screen "tryb_manualny" 800x480
   on GenerateScreen: SetTag("Tag_ScreenNumber", 2)
   TextField "Text field_1" at 282,4 size 223x34; Text 'TRYB MANUALNY'
   TextField "Text field_4" at 512,155 size 171x61; Text 'STOPIEŃ OTWARCIA OKIEN OTWIERANIE OKIEN'
   Button "Button_4" at 518,261 size 80x70; TextOff 'PODLEWANIE'
      on Click: InvertBit("Przycisk_podlewania_manual")
   Button "Button_5" at 611,261 size 80x70; TextOff 'GRZANIE'
      on Click: InvertBit("Przycisk_grzanie_manual")
   Button "Button_6" at 701,261 size 80x70; TextOff 'WENTYLACJA'
      on Click: InvertBit("Przycisk_wentylacja_manual")
   GraphicView "Graphic view_1" at 710,356 size 60x60; Picture "fan_4829316"
      Visibility <- "Wentylator"
   GraphicView "Graphic view_6" at 622,356 size 60x60; Picture "heater_4463010"
      Visibility <- "Grzałka"
   GraphicView "Graphic view_7" at 527,356 size 64x60; Picture "irrigation_18631825"
      Visibility <- "Pompa_podlewanie"
   GraphicView "Graphic view_9" at 710,356 size 60x60; Picture "fan_off"
      Visibility <- "Wentylator"
   GraphicView "Graphic view_10" at 622,356 size 60x60; Picture "heater_off"
      Visibility <- "Grzałka"
   GraphicView "Graphic view_11" at 527,356 size 64x60; Picture "irrigation_off"
      Visibility <- "Pompa_podlewanie"
   Button "Button_14" at 3,1 size 43x43; TextOff 'DOM'; PictureOff "home_1"
      on Click: ActivateScreen("Root screen", 0)
   Button "Button_1" at 750,0 size 50x50; TextOff 'Text'; PictureOff "Back_arrow"
      on Click: function_efd93a16()
   Circle "Circle_1" at 541,428 size 42x42
      Visibility <- "Pompa_podlewanie"
   Circle "Circle_4" at 541,428 size 42x42
      Visibility <- "Pompa_podlewanie"
   Circle "Circle_2" at 631,428 size 42x42
      Visibility <- "Grzałka"
   Circle "Circle_5" at 631,428 size 42x42
      Visibility <- "Grzałka"
   Circle "Circle_3" at 720,428 size 41x41
      Visibility <- "Wentylator"
   Circle "Circle_6" at 720,428 size 41x41
      Visibility <- "Wentylator"
   TextField "Text field_8" at 405,71 size 117x61; Text 'STOPIEŃ OTWARCIA OKIEN STOPIEŃ ZASŁONIECIA ROLET'
   Bar "Bar_6" at 625,71 size 165x66; MinimumValue 0; MaximumValue 100
      ProcessValue <- "Stopien_zasloniecia_rolet_manual"
   Button "Button_3" at 532,109 size 80x50; TextOff '+ / ODSŁOŃ'
      on Click: function_b9b71300("Stopien_zasloniecia_rolet_manual", 5)
   Button "Button_7" at 530,49 size 80x50; TextOff '- / ZASŁOŃ'
      on Press: function_dd21b452("Stopien_zasloniecia_rolet_manual", 5)
   Button "Button_2" at 425,261 size 80x70; TextOff 'PODLEWANIE / MIKROZRASZANIE'
      on Click: InvertBit("Przycisk_zraszania_manual")
   GraphicView "Graphic view_2" at 434,356 size 60x60; Picture "sprinkler_4552152"
      Visibility <- "Pompa_zraszacze"
   GraphicView "Graphic view_3" at 434,356 size 60x60; Picture "sprinkler"
      Visibility <- "Pompa_zraszacze"
   Circle "Circle_7" at 443,428 size 42x42
      Visibility <- "Pompa_zraszacze"
   Circle "Circle_8" at 443,428 size 42x42
      Visibility <- "Pompa_zraszacze"
   Switch "Switch_1" at 499,199 size 209x37; CaptionText 'Switch'; TextOff 'ZAMKNIĘTE'; TextOn 'OTWARTE'
      ProcessValue <- "Otwarcie_okien_man"
   TextField "Text field_3" at 10,365 size 166x23; Text 'SZYBKOŚĆ WIATRU'
   IOField "I/O field_3" at 61,397 size 70x65; FormatPattern 999
      ProcessValue <- "Czujnik_wiatru"
   IOField "I/O field_1" at 47,179 size 101x32; FormatPattern 99999
      ProcessValue <- "Czujnik_natezenia_światła"
   TextField "Text field_15" at 128,398 size 52x72; Text 'Km h'
   IOField "I/O field_2" at 43,282 size 83x65; FormatPattern 9999
      ProcessValue <- "Wewnetrzny_czujnik_CO2"
   TextField "Text field_11" at 117,291 size 69x39; Text 'ppm'
   TextField "Text field_5" at 13,138 size 204x23; Text 'INSOLATION / NASŁONECZNIENIE / SONNENEINSTRAHLUNG'
   IOField "I/O field_8" at 57,85 size 93x40; FormatPattern 99.99
      ProcessValue <- "Temperatura_wewnetrzna"
   TextField "Text field_20" at 26,42 size 137x42; Text 'TEMPERATURA TEMPERATURA WEWNTĘTRZNA'
   TextField "Text field_7" at 199,365 size 175x23; Text 'WILGOTNOŚĆ GLEBY'
   IOField "I/O field_5" at 247,283 size 83x65; FormatPattern 9999
      ProcessValue <- "Zewnetrzny_czujnik_CO2"
   IOField "I/O field_4" at 265,164 size 69x65; FormatPattern 999
      ProcessValue <- "Czujnik_wilgotności_powietrza"
   IOField "I/O field_6" at 260,395 size 68x65; FormatPattern 999
      ProcessValue <- "Czujnik_wilgotności_gleby"
   TextField "Text field_12" at 323,172 size 47x46; Text '%'
   TextField "Text field_13" at 320,406 size 47x46; Text '%'
   TextField "Text field_16" at 326,292 size 69x39; Text 'ppm'
   IOField "I/O field_9" at 247,75 size 97x65; FormatPattern 99.99
      ProcessValue <- "Temperatura_zewnetrzna"
   TextField "Text field_23" at 332,80 size 46x46; Text '°C'
   TextField "Text field_22" at 227,43 size 132x42; Text 'TEMPERATURA TEMPERATURA ZEWNĘTRZNA'
   TextField "Text field_9" at 228,246 size 123x42; Text 'STĘŻENIE CO2 ZEWNĘTRZNE STĘŻENIE CO2'
   TextField "Text field_6" at 180,137 size 223x42; Text 'WILGOTNOŚĆ POWIETRZA WILGOTNOŚĆ POWIETRZA'
   TextField "Text field_14" at 139,160 size 47x72; Text 'W m²'
   TextField "Text field_21" at 140,80 size 46x46; Text '°C'
   GraphicView "Graphic view_4" at 419,176 size 60x60; Picture "window_11250237"
   GraphicView "Graphic view_5" at 196,172 size 50x50; Picture "sensor_4212519"
   GraphicView "Graphic view_8" at 3,172 size 50x50; Picture "sensor_4212513"
   GraphicView "Graphic view_12" at 2,77 size 50x50; Picture "Thermometer_icon"
   GraphicView "Graphic view_13" at 198,77 size 50x50; Picture "Thermometer_icon"
   GraphicView "Graphic view_14" at 2,292 size 40x40; Picture "sensor_2828470"
   GraphicView "Graphic view_15" at 196,290 size 40x40; Picture "sensor_2828470"
   GraphicView "Graphic view_16" at 197,402 size 50x50; Picture "soil-sensor_11298794"
   GraphicView "Graphic view_17" at 2,406 size 50x50; Picture "anemometer_1113716"
   TextField "Text field_2" at 26,246 size 124x42; Text 'STĘŻENIE CO2 WEWNĘTRZNE STĘŻENIE CO2'

screen "praca" 800x480
   on GenerateScreen: SetTag("Tag_ScreenNumber", 5)
   GraphicView "Graphic view_4" at 274,396 size 70x70; Picture "soil-sensor_11298794"
   GraphicView "Graphic view_3" at 3,175 size 70x70; Picture "sensor_4212513"
   GraphicView "Graphic view_5" at 267,175 size 70x70; Picture "sensor_4212519"
   GraphicView "Graphic view_1" at 559,396 size 70x70; Picture "fan_4829316"
      Visibility <- "Wentylator"
   GraphicView "Graphic view_6" at 560,270 size 70x70; Picture "heater_4463010"
      Visibility <- "Grzałka"
   GraphicView "Graphic view_7" at 559,164 size 70x70; Picture "irrigation_18631825"
      Visibility <- "Pompa_podlewanie"
   GraphicView "Graphic view_8" at 11,397 size 70x70; Picture "anemometer_1113716"
   GraphicView "Graphic view_9" at 559,396 size 70x70; Picture "fan_off"
      Visibility <- "Wentylator"
   GraphicView "Graphic view_10" at 560,270 size 70x70; Picture "heater_off"
      Visibility <- "Grzałka"
   GraphicView "Graphic view_11" at 559,164 size 70x70; Picture "irrigation_off"
      Visibility <- "Pompa_podlewanie"
   GraphicView "Graphic view_12" at 278,267 size 70x70; Picture "sensor_2828470"
   TextField "Text field_1" at 52,152 size 204x23; Text 'INSOLATION / NASŁONECZNIENIE / SONNENEINSTRAHLUNG'
   TextField "Text field_3" at 44,373 size 166x23; Text 'SZYBKOŚĆ WIATRU'
   TextField "Text field_5" at 289,152 size 223x23; Text 'WILGOTNOŚĆ POWIETRZA'
   TextField "Text field_6" at 318,373 size 175x23; Text 'WILGOTNOŚĆ GLEBY'
   TextField "Text field_7" at 628,148 size 116x23; Text 'PODLEWANIE'
   TextField "Text field_8" at 638,252 size 80x23; Text 'GRZANIE'
   TextField "Text field_9" at 627,373 size 117x23; Text 'WENTYLACJA'
   TextField "Text field_10" at 81,3 size 256x34; Text 'PODGLĄD NA ŻYWO'
   Button "Button_1" at 750,0 size 50x50; TextOff 'WRÓĆ'; PictureOff "Back_arrow"
      on Click: function_efd93a16(); SetBit("HMI_Reset_Trybow")
   Button "Button_2" at 3,1 size 43x43; TextOff 'DOM'; PictureOff "home_1"
      on Click: ActivateScreen("Root screen", 0); SetBit("HMI_Reset_Trybow")
   IOField "I/O field_3" at 94,402 size 70x65; FormatPattern 999
      ProcessValue <- "Czujnik_wiatru"
   IOField "I/O field_5" at 348,277 size 83x65; FormatPattern 9999
      ProcessValue <- "Zewnetrzny_czujnik_CO2"
   IOField "I/O field_4" at 377,172 size 69x65; FormatPattern 999
      ProcessValue <- "Czujnik_wilgotności_powietrza"
   IOField "I/O field_6" at 381,397 size 68x65; FormatPattern 999
      ProcessValue <- "Czujnik_wilgotności_gleby"
   TextField "Text field_12" at 446,190 size 47x46; Text '%'
   TextField "Text field_13" at 466,405 size 47x46; Text '%'
   TextField "Text field_14" at 192,164 size 47x72; Text 'W m²'
   IOField "I/O field_1" at 83,190 size 101x32; FormatPattern 99999
      ProcessValue <- "Czujnik_natezenia_światła"
   TextField "Text field_15" at 173,402 size 52x72; Text 'Km h'
   Circle "Circle_1" at 703,188 size 48x48
      Visibility <- "Pompa_podlewanie"
   Circle "Circle_2" at 702,283 size 48x48
      Visibility <- "Grzałka"
   TextField "Text field_16" at 447,283 size 69x39; Text 'ppm'
   Circle "Circle_4" at 703,188 size 48x48
      Visibility <- "Pompa_podlewanie"
   Circle "Circle_5" at 702,283 size 48x48
      Visibility <- "Grzałka"
   Circle "Circle_3" at 703,415 size 48x48
      Visibility <- "Wentylator"
   Circle "Circle_6" at 703,415 size 48x48
      Visibility <- "Wentylator"
   TextField "Text field_17" at 381,3 size 288x34; Text 'PODGLĄD NA ŻYWO / TRYB AUTOMATYCZNY'
      Visibility <- "HMI_Aktywacja_trybu_automatycznego"
   GraphicView "Graphic view_13" at 560,63 size 70x70; Picture "sprinkler_4552152"
      Visibility <- "Pompa_zraszacze"
   GraphicView "Graphic view_14" at 560,63 size 70x70; Picture "sprinkler"
      Visibility <- "Pompa_zraszacze"
   Circle "Circle_7" at 703,83 size 48x48
      Visibility <- "Pompa_zraszacze"
   Circle "Circle_8" at 703,83 size 48x48
      Visibility <- "Pompa_zraszacze"
   TextField "Text field_19" at 609,44 size 156x23; Text 'PODLEWANIE / MIKROZRASZANIE'
   GraphicView "Graphic view_15" at 0,66 size 70x70; Picture "Thermometer_icon"
   IOField "I/O field_8" at 73,73 size 97x65; FormatPattern 99.99
      ProcessValue <- "Temperatura_wewnetrzna"
   TextField "Text field_21" at 171,85 size 46x46; Text '°C'
   GraphicView "Graphic view_16" at 275,66 size 70x70; Picture "Thermometer_icon"
   IOField "I/O field_9" at 348,73 size 97x65; FormatPattern 99.99
      ProcessValue <- "Temperatura_zewnetrzna"
   TextField "Text field_23" at 447,82 size 46x46; Text '°C'
   TextField "Text field_20" at 57,44 size 137x42; Text 'TEMPERATURA TEMPERATURA WEWNTĘTRZNA'
   TextField "Text field_22" at 334,44 size 132x42; Text 'TEMPERATURA TEMPERATURA ZEWNĘTRZNA'
   GraphicView "Graphic view_2" at 11,273 size 70x70; Picture "sensor_2828470"
   IOField "I/O field_2" at 81,283 size 83x65; FormatPattern 9999
      ProcessValue <- "Wewnetrzny_czujnik_CO2"
   TextField "Text field_11" at 180,289 size 69x39; Text 'ppm'
   TextField "Text field_2" at 83,252 size 124x42; Text 'STĘŻENIE CO2 WEWNĘTRZNE STĘŻENIE CO2'
   TextField "Text field_4" at 352,256 size 123x42; Text 'STĘŻENIE CO2 ZEWNĘTRZNE STĘŻENIE CO2'
   TextField "Text field_18" at 381,3 size 211x34; Text 'TRYB RECEPTUR'
      Visibility <- "HMI_Aktywacja_trybu_Receptur"

Template "Template_1" 800x480
   Button "Exit" at 671,429 size 71x50; TextOn 'Exit'; TextOff 'Exit'; PictureOn "ExitRuntime_KTP700_Basic_PN_TR"; PictureOff "ExitRuntime_KTP700_Basic_PN_TR"
      on Release: StopRuntime(0)
   Button "Alarms" at 524,429 size 71x50; TextOn 'Alarms'; TextOff 'Alarms'; PictureOn "AlarmDisplay_KTP700_Basic_PN_TR"; PictureOff "AlarmDisplay_KTP700_Basic_PN_TR"
      on Release: function_ef3f5d25("Alarm window_Unacknowledged", -1)
   Button "Start screen" at 169,429 size 71x50; TextOn 'Start screen'; TextOff 'Start screen'; PictureOn "NavigateHome_KTP700_Basic_PN_TR"; PictureOff "NavigateHome_KTP700_Basic_PN_TR"
      on Release: ActivateScreen("Root screen", 0)
      Visibility <- "AlwaysTRUE"
   Button "Language" at 377,429 size 71x50; TextOn 'Language'; TextOff 'Language'; PictureOn "ToggleLanguage_KTP700_Basic_PN_TR"; PictureOff "ToggleLanguage_KTP700_Basic_PN_TR"
      on Release: function_fb9197e8(-1)

screen "Receptury" 800x480
   RecipeView "Recipe view_1" at 0,38 size 799x413; Recipe "Receptura_nr1"; RecipeNameCaption 'Recipe Name: / Wybierz Recepturę / Rezepturname:'; EntryNameCaption 'Entry Name / Zapisane Parametry / Eintragsname'; DataRecordNameCaption 'Data Record Name: / Wybierz Recepturę / Datensatzname:'
   GraphicView "Graphic view_1" at 529,152 size 35x35; Picture "Thermometer_icon"
   GraphicView "Graphic view_2" at 529,190 size 35x35; Picture "sensor_4212519"
   GraphicView "Graphic view_3" at 529,230 size 35x35; Picture "soil-sensor_11298794"
   GraphicView "Graphic view_4" at 529,269 size 35x35; Picture "window_11250237"
   GraphicView "Graphic view_5" at 529,308 size 35x35; Picture "sensor_2828470"
   GraphicView "Graphic view_6" at 529,348 size 35x35; Picture "sensor_4212513"
   TextField "Text field_11" at 569,150 size 39x38; Text '°C'
   TextField "Text field_18" at 569,190 size 39x38; Text '%'
   TextField "Text field_1" at 569,230 size 39x38; Text '%'
   TextField "Text field_2" at 564,269 size 57x32; Text '1/0'
   TextField "Text field_16" at 563,308 size 55x32; Text 'ppm'
   TextField "Text field_6" at 576,339 size 28x50; Text '°C W m'
   TextField "Text field_3" at 593,362 size 31x17; Text '2'
   Button "Button_1" at 750,0 size 50x50; TextOff 'WRÓĆ'; PictureOff "Back_arrow"
      on Click: function_efd93a16()
   Button "Button_14" at 3,1 size 43x43; TextOff 'DOM'; PictureOff "home_1"
      on Click: ActivateScreen("Root screen", 0)
   TextField "Text field_4" at 320,2 size 170x37; Text 'RECEPTURY'
   TextField "Text field_5" at 12,448 size 50x23; Text 'Nowy'
   TextField "Text field_7" at 69,448 size 57x23; Text 'Zapisz'
   TextField "Text field_8" at 137,448 size 45x23; Text 'Usuń'
   TextField "Text field_9" at 190,438 size 60x42; Text 'Zmień Nazwę'
   TextField "Text field_10" at 663,438 size 66x42; Text 'Załaduj z PLC'
   TextField "Text field_12" at 729,438 size 66x42; Text 'Załaduj do PLC'
   Button "Button_2" at 405,402 size 255x40; TextOff 'ZATWIERDŹ'
      on Click: ResetBit("HMI_Reset_Trybow"); ActivateScreen("praca", 0); SetBit("HMI_Aktywacja_trybu_Receptur")
   TextField "Text field_13" at 456,450 size 173x23; Text 'Przejdź w tryb pracy'
   Button "Button_3" at 256,401 size 140x40; TextOff 'Z'
      on Click: function_ea909784(1, U 0, '\USB_X60.1\record.csv', 2, 1, N)
   TextField "Text field_14" at 266,438 size 113x42; Text 'Zapisz Kopię zapasową'

screen "Symulacja_czujnikow" 800x480
   TextField "Text field_1" at 21,47 size 252x23; Text 'Czujnik Wilgotności powietrza'
   TextField "Text field_2" at 308,47 size 214x23; Text 'Czujnik Wilgotności gleby'
   TextField "Text field_3" at 32,202 size 202x23; Text 'Termometr wewnętrzny'
   TextField "Text field_4" at 323,202 size 197x23; Text 'Termometr zewnętrzny'
   TextField "Text field_5" at 569,47 size 216x23; Text 'Czujnik natężenia światła'
   TextField "Text field_6" at 607,202 size 124x23; Text 'Czujnik wiatru'
   TextField "Text field_7" at 27,346 size 208x23; Text 'Wewnętrzny czujnik CO2'
   TextField "Text field_8" at 306,346 size 202x23; Text 'Zewnętrzny czujnik CO2'
   TextField "Text field_9" at 569,346 size 206x23; Text 'Stopień zasłonięcia rolet'
   IOField "I/O field_4" at 599,83 size 150x60; FormatPattern 9999
      ProcessValue <- "Czujnik_natezenia_światła"
   IOField "I/O field_5" at 599,242 size 150x60; FormatPattern 999
      ProcessValue <- "Czujnik_wiatru"
   IOField "I/O field_6" at 69,375 size 150x60; FormatPattern 9999
      ProcessValue <- "Wewnetrzny_czujnik_CO2"
   IOField "I/O field_7" at 346,375 size 150x60; FormatPattern 9999
      ProcessValue <- "Zewnetrzny_czujnik_CO2"
   IOField "I/O field_8" at 599,375 size 150x60; FormatPattern 999
      ProcessValue <- "Stopien_zasloniecia_rolet"
   IOField "I/O field_10" at 69,83 size 150x60; FormatPattern 999
      ProcessValue <- "Czujnik_wilgotności_powietrza"
   IOField "I/O field_11" at 346,83 size 150x60; FormatPattern 999
      ProcessValue <- "Czujnik_wilgotności_gleby"
   IOField "I/O field_12" at 69,242 size 150x60; FormatPattern 99.9
      ProcessValue <- "Temperatura_wewnetrzna"
   IOField "I/O field_13" at 346,242 size 150x60; FormatPattern 99.9
      ProcessValue <- "Temperatura_zewnetrzna"
   TextField "Text field_10" at 248,5 size 321x34; Text 'ZAPISZ RECEPTURE / SYMULACJA CZUJNIKÓW'
   Button "Button_1" at 750,0 size 50x50; TextOff 'WRÓĆ'; PictureOff "Back_arrow"
      on Click: function_efd93a16()
   Button "Button_14" at 3,1 size 43x43; TextOff 'DOM'; PictureOff "home_1"
      on Click: ActivateScreen("Root screen", 0)

screen "tryb_automatyczny" 800x480
   on GenerateScreen: SetTag("Tag_ScreenNumber", 1)
   IOField "I/O field_1" at 67,301 size 57x40; FormatPattern 99.9
      ProcessValue <- "Temperatura_wewnetrzna"
   Button "Button_1" at 750,0 size 50x50; TextOff 'WRÓĆ'; PictureOff "Back_arrow"
      on Click: function_efd93a16()
   Button "Button_2" at 530,382 size 259x89; TextOff 'ZATWIERDŹ'
      on Click: ResetBit("HMI_Reset_Trybow"); SetBit("HMI_Aktywacja_trybu_automatycznego"); ActivateScreen("praca", 0)
   Bar "Bar_1" at 7,89 size 50x250; MinimumValue 0; MaximumValue 45
      ProcessValue <- "Temperatura_auto"
   TextField "Text field_2" at 1,50 size 132x23; Text 'TEMPERATURA'
   Bar "Bar_2" at 170,90 size 50x250; MinimumValue 0; MaximumValue 100
      ProcessValue <- "Wilgotnosc_powietrza_auto"
   TextField "Text field_3" at 165,47 size 122x42; Text 'WOLGOTNOŚĆ POWIETRZA WILGOTNOŚĆ POWIETRZA'
   Button "Button_3" at 71,94 size 75x45; TextOff '+ / +0.5 °C'
      on Press: function_dd21b452("Temperatura_auto", 0.5)
   Button "Button_7" at 71,162 size 75x45; TextOff '- / -0.5 °C'
      on Press: function_b9b71300("Temperatura_auto", 0.5)
   IOField "I/O field_2" at 67,230 size 62x40; FormatPattern 99.9
      ProcessValue <- "Temperatura_auto"
   TextField "Text field_11" at 122,239 size 23x22; Text '°C'
   TextField "Text field_9" at 122,312 size 23x22; Text '°C'
   Bar "Bar_4" at 335,90 size 50x250; MinimumValue 0; MaximumValue 100
      ProcessValue <- "Wilgotnosc_gleby_auto"
   TextField "Text field_10" at 327,46 size 122x42; Text 'WOLGOTNOŚĆ GLEBY WILGOTNOŚĆ GLEBY'
   Button "Button_8" at 398,111 size 65x40; TextOff '+ / +2%'
      on Click: function_dd21b452("Wilgotnosc_gleby_auto", 2)
   Button "Button_9" at 398,160 size 65x40; TextOff '- / -2%'
      on Click: function_b9b71300("Wilgotnosc_gleby_auto", 2)
   IOField "I/O field_5" at 402,234 size 60x40; FormatPattern 999
      ProcessValue <- "Wilgotnosc_gleby_auto"
   IOField "I/O field_6" at 404,304 size 58x40; FormatPattern 999
      ProcessValue <- "Czujnik_wilgotności_gleby"
   TextField "Text field_12" at 385,222 size 101x22; Text 'USTAWIONA'
   TextField "Text field_13" at 389,293 size 86x22; Text 'AKTUALNA'
   TextField "Text field_14" at 439,243 size 23x22; Text '%'
   TextField "Text field_15" at 439,314 size 23x22; Text '%'
   Button "Button_10" at 229,105 size 65x40; TextOff '+ / +5%'
      on Click: function_dd21b452("Wilgotnosc_powietrza_auto", 5)
   Button "Button_11" at 229,165 size 65x40; TextOff '- / -5%'
      on Click: function_b9b71300("Wilgotnosc_powietrza_auto", 5)
   IOField "I/O field_4" at 234,227 size 66x40; FormatPattern 999
      ProcessValue <- "Wilgotnosc_powietrza_auto"
   IOField "I/O field_7" at 236,299 size 62x40; FormatPattern 999
      ProcessValue <- "Czujnik_wilgotności_powietrza"
   TextField "Text field_16" at 223,214 size 101x22; Text 'USTAWIONA'
   TextField "Text field_17" at 223,285 size 86x22; Text 'AKTUALNA'
   TextField "Text field_18" at 275,236 size 23x22; Text '%'
   TextField "Text field_19" at 275,307 size 23x22; Text '%'
   Button "Button_14" at 3,1 size 43x43; TextOff 'DOM'; PictureOff "home_1"
      on Click: ActivateScreen("Root screen", 0)
   TextField "Text field_4" at 124,384 size 128x23; Text 'SYSTEM OKIEN'
   Switch "Switch_1" at 106,410 size 181x46; TextOn 'ON'; CaptionText 'Switch'; TextOff 'OFF'
      ProcessValue <- "System_okien_auto"
   GraphicView "Graphic view_1" at 128,46 size 40x40; Picture "Thermometer_icon"
   GraphicView "Graphic view_2" at 281,47 size 40x40; Picture "sensor_4212519"
   TextField "Text field_5" at 60,288 size 86x22; Text 'AKTUALNA'
   TextField "Text field_6" at 57,216 size 101x22; Text 'USTAWIONA'
   GraphicView "Graphic view_3" at 443,50 size 40x40; Picture "soil-sensor_11298794"
   TextField "Text field_1" at 250,4 size 288x34; Text 'TRYB AUTOMATYCZNY'
   Bar "Bar_3" at 496,90 size 50x250; MinimumValue 0; MaximumValue 1500
      ProcessValue <- "Naslonecznienie_auto"
   TextField "Text field_7" at 487,38 size 154x40; Text 'WOLGOTNOŚĆ GLEBY NASŁONECZNIENIE'
   GraphicView "Graphic view_4" at 585,65 size 40x40; Picture "sensor_4212513"
   Button "Button_4" at 553,110 size 82x43; TextOff '+ +50 W m'
      on Click: function_dd21b452("Naslonecznienie_auto", 50)
   Button "Button_5" at 554,165 size 82x43; TextOff '- -50 W m'
      on Click: function_b9b71300("Naslonecznienie_auto", 50)
   IOField "I/O field_3" at 561,233 size 61x40; FormatPattern 9999
      ProcessValue <- "Naslonecznienie_auto"
   TextField "Text field_8" at 545,221 size 101x22; Text 'USTAWIONA / USTAWIONE'
   IOField "I/O field_8" at 563,304 size 62x40; FormatPattern 9999
      ProcessValue <- "Czujnik_natezenia_światła"
   TextField "Text field_20" at 549,292 size 86x22; Text 'AKTUALNA / AKTUALNE'
   TextField "Text field_23" at 616,129 size 32x18; Text '2'
   TextField "Text field_24" at 614,184 size 32x18; Text '2'
   Bar "Bar_5" at 656,90 size 45x250; MinimumValue 400; MaximumValue 950
      ProcessValue <- "Poziom_CO2_auto"
   TextField "Text field_21" at 650,47 size 128x23; Text 'SYSTEM OKIEN / POZIOM CO2'
   IOField "I/O field_9" at 723,233 size 66x40; FormatPattern 999
      ProcessValue <- "Poziom_CO2_auto"
   TextField "Text field_22" at 699,216 size 101x22; Text 'USTAWIONA / USTAWIONE'
   IOField "I/O field_10" at 723,312 size 62x40; FormatPattern 999
      ProcessValue <- "Wewnetrzny_czujnik_CO2"
   TextField "Text field_25" at 708,293 size 86x22; Text 'AKTUALNA'
   Button "Button_6" at 714,113 size 73x40; TextOff '+ / +25ppm'
      on Click: function_dd21b452("Poziom_CO2_auto", 25)
   Button "Button_12" at 714,165 size 73x40; TextOff '+ / -25ppm'
      on Click: function_b9b71300("Poziom_CO2_auto", 25)
   GraphicView "Graphic view_5" at 754,54 size 40x40; Picture "sensor_2828470"
   GraphicView "Graphic view_6" at 17,400 size 55x55; Picture "window_11250237"
   TextField "Text field_26" at 339,400 size 164x42; Text 'miejsce na ewentualne zmiany'
*)